(* Logix 5000 project; controller NWGG 1756-L72 rev 35.12; software revision 35.00; part 6 of 19 *)
(* tags used below, declared in another part *)
   _124MB : ALIAS FOR B9[124].2;
   _124STB : ALIAS FOR B9[124].0;
   _124STPB : ALIAS FOR B9[124].1;
   _24_16_0 : ALIAS FOR N250[0];
   _24_16_1 : ALIAS FOR N250[1];
   _24_16_2 : ALIAS FOR N250[2];
   _24_16_3 : ALIAS FOR N250[3];
   _24_16_4 : ALIAS FOR N250[4];
   _24_16_5 : ALIAS FOR N250[5];
   _24_16_6 : ALIAS FOR N250[6];
   _24_16_7 : ALIAS FOR N250[7];
   _24_17_0 : ALIAS FOR N240[0];
   _24_18_0_AN : ALIAS FOR N230[10];
   _24_18_1_AN : ALIAS FOR N230[11];
   _24_18_2_AN : ALIAS FOR N230[12];
   _24_18_3_AN : ALIAS FOR N230[13];
   _24_19_0 : ALIAS FOR N220[10];
   _24_19_1 : ALIAS FOR N220[11];
   _24_19_2 : ALIAS FOR N220[12];
   _24_19_3 : ALIAS FOR N220[13];
   _24_20_0 : ALIAS FOR N210[10];
   _45_AIR_SEQ : ALIAS FOR T4[34];
   _45_SEQ_AIR : ALIAS FOR O12.15;
   _45AUTO : ALIAS FOR B9[45].4;
   _45HAND : ALIAS FOR B9[45].3;
   _45M : ALIAS FOR O25[8].7;
   _45MB : ALIAS FOR B9[45].2;
   _45STB : ALIAS FOR B9[45].0;
   _45STPB : ALIAS FOR B9[45].1;
   _45Y : ALIAS FOR I25[0].7;
   _46AUTO : ALIAS FOR B9[46].4;
   _46HAND : ALIAS FOR B9[46].3;
   _46M : ALIAS FOR O25[8].8;
   _46MB : ALIAS FOR B9[46].2;
   _46STB : ALIAS FOR B9[46].0;
   _46STPB : ALIAS FOR B9[46].1;
   _46Y : ALIAS FOR I25[0].8;
   _47M : ALIAS FOR O25[9].10;
   _47MB : ALIAS FOR B9[47].2;
   _47Y : ALIAS FOR I25[1].10;
   _700_TREAT : ALIAS FOR I7.3;
   _9_TRT_MOV : ALIAS FOR O24[7].4;
   ALARM_FIEL : ALIAS FOR T11[7];
   ALARM_HAND : ALIAS FOR B3[0].10;
   ALARM_HORN : ALIAS FOR O25[11].15;
   ALARM_HORN1 : ALIAS FOR O12.14;
   ALARM_LIGH : ALIAS FOR O13.15;
   ALARM_LT_O : ALIAS FOR T11[3];
   ALARM_SILE : ALIAS FOR I25[4].7;
   ALARM_SILE1 : ALIAS FOR I7.13;
   ALARM_SILE2 : ALIAS FOR B3[0].3;
   ALARM_SILE4 : ALIAS FOR B3[0].9;
   ALRM_LIGHT : ALIAS FOR O25[11].14;
   ALRM_SILEN : ALIAS FOR B3[0].7;
   B3 : DINT[250];
   I24_004_Bit00 : ALIAS FOR I24[4].0;
   I24_004_Bit01 : ALIAS FOR I24[4].1;
   I24_004_Bit02 : ALIAS FOR I24[4].2;
   I24_004_Bit03 : ALIAS FOR I24[4].3;
   I24_004_Bit04 : ALIAS FOR I24[4].4;
   I24_004_Bit05 : ALIAS FOR I24[4].5;
   I24_004_Bit06 : ALIAS FOR I24[4].6;
   I24_004_Bit07 : ALIAS FOR I24[4].7;
   I24_004_Bit08 : ALIAS FOR I24[4].8;
   I24_006_Bit02 : ALIAS FOR I24[6].2;
   I24_021_Bit00 : ALIAS FOR I24[21].0;
   I24_021_Bit01 : ALIAS FOR I24[21].1;
   I24_021_Bit02 : ALIAS FOR I24[21].2;
   I24_021_Bit03 : ALIAS FOR I24[21].3;
   I24_021_Bit04 : ALIAS FOR I24[21].4;
   I24_021_Bit05 : ALIAS FOR I24[21].5;
   I24_021_Bit06 : ALIAS FOR I24[21].6;
   I24_021_Bit07 : ALIAS FOR I24[21].7;
   I24_021_Bit08 : ALIAS FOR I24[21].8;
   IE8_BTR_FL : ALIAS FOR N23[0];
   MAIN_TIMER1 : ALIAS FOR T11[1];
   N23 : DINT[5];
   O24_005_Bit15 : ALIAS FOR O24[5].15;
   O24_007_Bit10 : ALIAS FOR O24[7].10;
   P10_FLOW_A : ALIAS FOR N13[82];
   P10_FLOW_P1 : ALIAS FOR C5[39];
   P10_FLW_OZ : ALIAS FOR N13[80];
   P10_MB : ALIAS FOR B12[10].2;
   P10_OZ : ALIAS FOR N13[81];
   P10_SET : ALIAS FOR B12[10].0;
   P10_SPEED : ALIAS FOR N13[84];
   P10_STOP : ALIAS FOR B12[10].1;
   P1_FLOW_AN : ALIAS FOR N13[2];
   P1_FLOW_PL : ALIAS FOR C5[30];
   P1_FLW_OZ : ALIAS FOR N13[0];
   P1_MB : ALIAS FOR B12[1].2;
   P1_OZ : ALIAS FOR N13[1];
   P1_SET : ALIAS FOR B12[1].0;
   P1_SPEED_O : ALIAS FOR N13[4];
   P1_STOP : ALIAS FOR B12[1].1;
   P2_FLOW_AN : ALIAS FOR N13[12];
   P2_FLOW_PL : ALIAS FOR C5[32];
   P2_FLW_OZ : ALIAS FOR N13[10];
   P2_MB : ALIAS FOR B12[2].2;
   P2_OZ : ALIAS FOR N13[11];
   P2_SET : ALIAS FOR B12[2].0;
   P2_SPEED_O : ALIAS FOR N13[14];
   P2_STOP : ALIAS FOR B12[2].1;
   P3_FLOW_AN : ALIAS FOR N13[22];
   P3_FLOW_PL : ALIAS FOR C5[33];
   P3_FLW_OZ : ALIAS FOR N13[20];
   P3_MB : ALIAS FOR B12[3].2;
   P3_OZ : ALIAS FOR N13[21];
   P3_SET : ALIAS FOR B12[3].0;
   P3_SPEED_O : ALIAS FOR N13[24];
   P3_STOP : ALIAS FOR B12[3].1;
   P4_FLOW_AN : ALIAS FOR N13[32];
   P4_FLOW_PL : ALIAS FOR C5[34];
   P4_FLW_OZ : ALIAS FOR N13[30];
   P4_MB : ALIAS FOR B12[4].2;
   P4_OZ : ALIAS FOR N13[31];
   P4_SET : ALIAS FOR B12[4].0;
   P4_SPEED_O : ALIAS FOR N13[34];
   P4_STOP : ALIAS FOR B12[4].1;
   P5_FLOW_AN : ALIAS FOR N13[42];
   P5_FLOW_PL : ALIAS FOR C5[35];
   P5_FLW_OZ : ALIAS FOR N13[40];
   P5_MB : ALIAS FOR B12[5].2;
   P5_OZ : ALIAS FOR N13[41];
   P5_SET : ALIAS FOR B12[5].0;
   P5_SPEED_O : ALIAS FOR N13[44];
   P5_STOP : ALIAS FOR B12[5].1;
   P6_FLOW_AN : ALIAS FOR N13[52];
   P6_FLOW_PL : ALIAS FOR C5[36];
   P6_FLW_OZ : ALIAS FOR N13[50];
   P6_MB : ALIAS FOR B12[6].2;
   P6_OZ : ALIAS FOR N13[51];
   P6_SET : ALIAS FOR B12[6].0;
   P6_SPEED_O : ALIAS FOR N13[54];
   P6_STOP : ALIAS FOR B12[6].1;
   P7_FLOW_AN : ALIAS FOR N13[62];
   P7_FLOW_PL : ALIAS FOR C5[37];
   P7_FLW_OZ : ALIAS FOR N13[60];
   P7_MB : ALIAS FOR B12[7].2;
   P7_OZ : ALIAS FOR N13[61];
   P7_SET : ALIAS FOR B12[7].0;
   P7_SPEED_O : ALIAS FOR N13[64];
   P7_STOP : ALIAS FOR B12[7].1;
   P8_FLOW_AN : ALIAS FOR N13[72];
   P8_FLOW_PL : ALIAS FOR C5[38];
   P8_FLW_OZ : ALIAS FOR N13[70];
   P8_MB : ALIAS FOR B12[8].2;
   P8_OZ : ALIAS FOR N13[71];
   P8_SET : ALIAS FOR B12[8].0;
   P8_SPEED_O : ALIAS FOR N13[74];
   P8_STOP : ALIAS FOR B12[8].1;
   P_RESET_AU : ALIAS FOR B3[4].0;
   RSVIEW_ALA : ALIAS FOR B3[0].11;
   T11_DLY_TR : ALIAS FOR T4[0].PRE;
   T11_DLY_TR2 : ALIAS FOR T4[1].PRE;
   T11_SET_DE : ALIAS FOR B3[2].0;
   T11_TREAT : ALIAS FOR B3[11].0;
   T11_TRT_MO1 : ALIAS FOR T4[41].PRE;
   T12_DLY_TR1 : ALIAS FOR T4[2].PRE;
   T12_DLY_TR4 : ALIAS FOR T4[3].PRE;
   T12_SET_DE : ALIAS FOR B3[2].1;
   T12_TREAT : ALIAS FOR B3[12].0;
   T12_TRT_MO1 : ALIAS FOR T4[42].PRE;
   T13_DLY_TR1 : ALIAS FOR T4[4].PRE;
   T13_DLY_TR4 : ALIAS FOR T4[5].PRE;
   T13_SET_DE : ALIAS FOR B3[2].2;
   T13_TREAT : ALIAS FOR B3[13].0;
   T13_TRT_MO1 : ALIAS FOR T4[43].PRE;
   T13C_CLOSE1 : ALIAS FOR T22[6].PRE;
   T13C_SET_D : ALIAS FOR B21[70].14;
   T13C_TRT_M1 : ALIAS FOR T22[7].PRE;
   T13C_TRT_O1 : ALIAS FOR T22[5].PRE;
   T14_DLY_TR2 : ALIAS FOR T4[6].ACC;
   T14_DLY_TR4 : ALIAS FOR T4[7].PRE;
   T14_SET_DE : ALIAS FOR B3[2].3;
   T14_TREAT : ALIAS FOR B3[14].0;
   T14_TRT_MO1 : ALIAS FOR T4[44].PRE;
   T15_SET_DE : ALIAS FOR B3[2].4;
   T15_TREAT : ALIAS FOR B3[15].0;
   T15_TRT_MO1 : ALIAS FOR T4[45].PRE;
   T15_TRT_OF1 : ALIAS FOR T4[9].PRE;
   T15_TRT_ON1 : ALIAS FOR T4[8].PRE;
   T16_SET_DE : ALIAS FOR B3[2].5;
   T16_TREAT : ALIAS FOR B3[16].0;
   T16_TRT_MO1 : ALIAS FOR T4[46].PRE;
   T16_TRT_OF1 : ALIAS FOR T4[11].PRE;
   T16_TRT_ON1 : ALIAS FOR T4[10].PRE;
   T17_SET_DE : ALIAS FOR B3[2].6;
   T17_TREAT : ALIAS FOR B3[17].0;
   T17_TRT_MO1 : ALIAS FOR T4[47].PRE;
   T17_TRT_OF1 : ALIAS FOR T4[13].PRE;
   T17_TRT_ON1 : ALIAS FOR T4[12].PRE;
   T19 : TIMER[2];
   T19C_CLOSE2 : ALIAS FOR T22[3].PRE;
   T19C_SET_D : ALIAS FOR B21[71].14;
   T19C_TRT_M1 : ALIAS FOR T22[4].PRE;
   T19C_TRT_O1 : ALIAS FOR T22[0].PRE;
   T21_SET_DE : ALIAS FOR B3[2].7;
   T21_TREAT : ALIAS FOR B3[21].0;
   T21_TRT_MO1 : ALIAS FOR T4[48].PRE;
   T21_TRT_OF1 : ALIAS FOR T4[15].PRE;
   T21_TRT_ON1 : ALIAS FOR T4[14].PRE;
   T22_SET_DE : ALIAS FOR B3[2].8;
   T22_TREAT : ALIAS FOR B3[22].0;
   T22_TRT_MO1 : ALIAS FOR T4[49].PRE;
   T22_TRT_OF1 : ALIAS FOR T4[17].PRE;
   T22_TRT_ON1 : ALIAS FOR T4[16].PRE;
   T23_SET_DE : ALIAS FOR B3[2].9;
   T23_TREAT : ALIAS FOR B3[23].0;
   T23_TRT_MO1 : ALIAS FOR T4[50].PRE;
   T23_TRT_OF1 : ALIAS FOR T4[19].PRE;
   T23_TRT_ON1 : ALIAS FOR T4[18].PRE;
   T24_SET_DE : ALIAS FOR B3[2].10;
   T24_TREAT : ALIAS FOR B3[24].0;
   T24_TRT_MO1 : ALIAS FOR T4[51].PRE;
   T24_TRT_OF1 : ALIAS FOR T4[21].PRE;
   T24_TRT_ON1 : ALIAS FOR T4[20].PRE;
   T25_SET_DE : ALIAS FOR B3[2].11;
   T25_TREAT : ALIAS FOR B3[25].0;
   T25_TRT_MO1 : ALIAS FOR T4[52].PRE;
   T25_TRT_OF1 : ALIAS FOR T4[23].PRE;
   T25_TRT_ON1 : ALIAS FOR T4[22].PRE;
   T26_SET_DE : ALIAS FOR B3[2].12;
   T26_TREAT : ALIAS FOR B3[26].0;
   T26_TRT_MO1 : ALIAS FOR T4[53].PRE;
   T26_TRT_OF1 : ALIAS FOR T4[25].PRE;
   T26_TRT_ON1 : ALIAS FOR T4[24].PRE;
   T27_SET_DE : ALIAS FOR B3[2].13;
   T27_TREAT : ALIAS FOR B3[27].0;
   T27_TRT_MO1 : ALIAS FOR T4[54].PRE;
   T27_TRT_OF1 : ALIAS FOR T4[27].PRE;
   T27_TRT_ON1 : ALIAS FOR T4[26].PRE;
   T28_SET_DE : ALIAS FOR B3[2].14;
   T28_TREAT : ALIAS FOR B3[28].0;
   T28_TRT_MO1 : ALIAS FOR T4[55].PRE;
   T28_TRT_OF1 : ALIAS FOR T4[29].PRE;
   T28_TRT_ON1 : ALIAS FOR T4[28].PRE;
   T29_SET_DE : ALIAS FOR B3[2].15;
   T29_TREAT : ALIAS FOR B3[29].0;
   T29_TRT_MO1 : ALIAS FOR T4[56].PRE;
   T29_TRT_OF1 : ALIAS FOR T4[31].PRE;
   T29_TRT_ON1 : ALIAS FOR T4[30].PRE;
   TRT_PumpRATE : DINT[50];
(* _2_MAIN, continued *)

ROUTINE _10_RAW_MOTORS   (* ladder *)
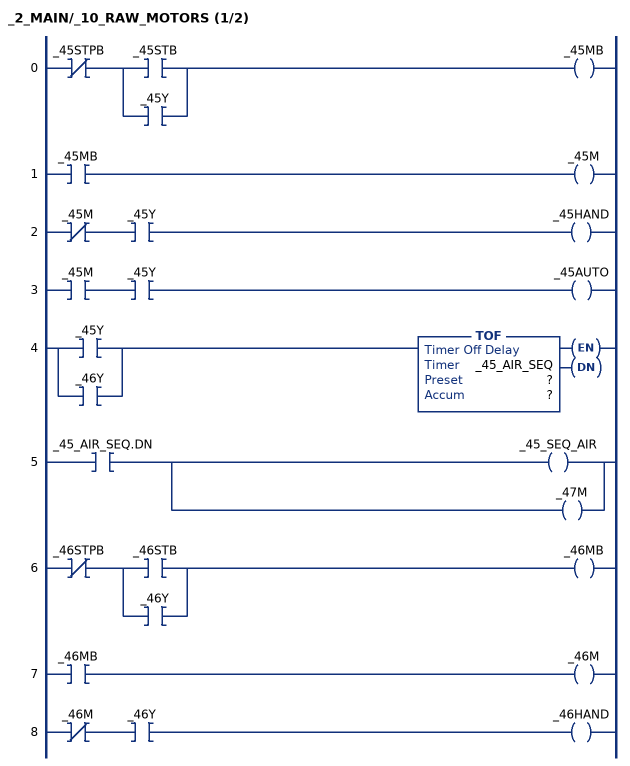
   0: XIO(_45STPB)[XIC(_45STB) ,XIC(_45Y) ]OTE(_45MB);
   1: XIC(_45MB)OTE(_45M);
   2: XIO(_45M)XIC(_45Y)OTE(_45HAND);
   3: XIC(_45M)XIC(_45Y)OTE(_45AUTO);
   4: [XIC(_45Y) ,XIC(_46Y) ]TOF(_45_AIR_SEQ,?,?);
   5: XIC(_45_AIR_SEQ.DN)[OTE(_45_SEQ_AIR) ,OTE(_47M) ];
   6: XIO(_46STPB)[XIC(_46STB) ,XIC(_46Y) ]OTE(_46MB);
   7: XIC(_46MB)OTE(_46M);
   8: XIO(_46M)XIC(_46Y)OTE(_46HAND);
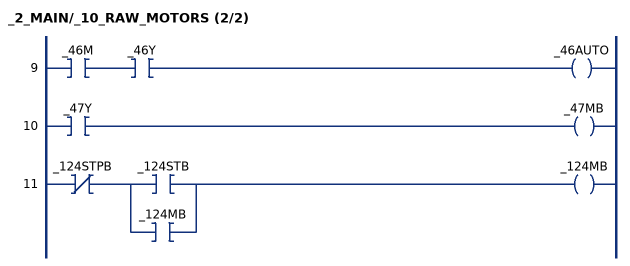
   9: XIC(_46M)XIC(_46Y)OTE(_46AUTO);
   10: XIC(_47Y)OTE(_47MB);
   11: XIO(_124STPB)[XIC(_124STB) ,XIC(_124MB) ]OTE(_124MB);
END_ROUTINE

ROUTINE _34_34_ALARMS   (* ladder *)
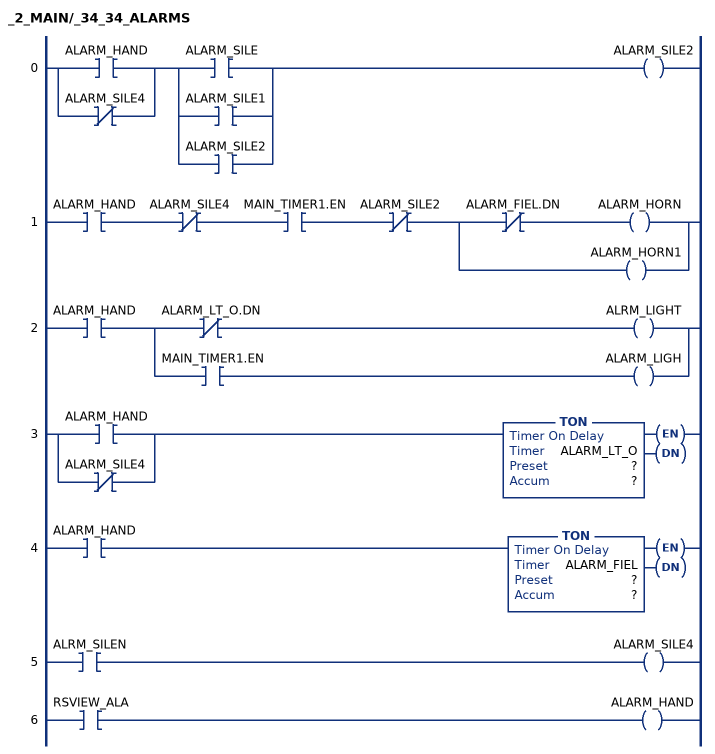
   0: [XIC(ALARM_HAND) ,XIO(ALARM_SILE4) ][XIC(ALARM_SILE) ,XIC(ALARM_SILE1) ,XIC(ALARM_SILE2) ]OTE(ALARM_SILE2);
   1: XIC(ALARM_HAND)XIO(ALARM_SILE4)XIC(MAIN_TIMER1.EN)XIO(ALARM_SILE2)[XIO(ALARM_FIEL.DN) OTE(ALARM_HORN) ,OTE(ALARM_HORN1) ];
   2: XIC(ALARM_HAND)[XIO(ALARM_LT_O.DN) OTE(ALRM_LIGHT) ,XIC(MAIN_TIMER1.EN) OTE(ALARM_LIGH) ];
   3: [XIC(ALARM_HAND) ,XIO(ALARM_SILE4) ]TON(ALARM_LT_O,?,?);
   4: XIC(ALARM_HAND)TON(ALARM_FIEL,?,?);
   5: XIC(ALRM_SILEN)OTE(ALARM_SILE4);
   6: XIC(RSVIEW_ALA)OTE(ALARM_HAND);
END_ROUTINE

ROUTINE _35_35_DEFAULT   (* ladder *)
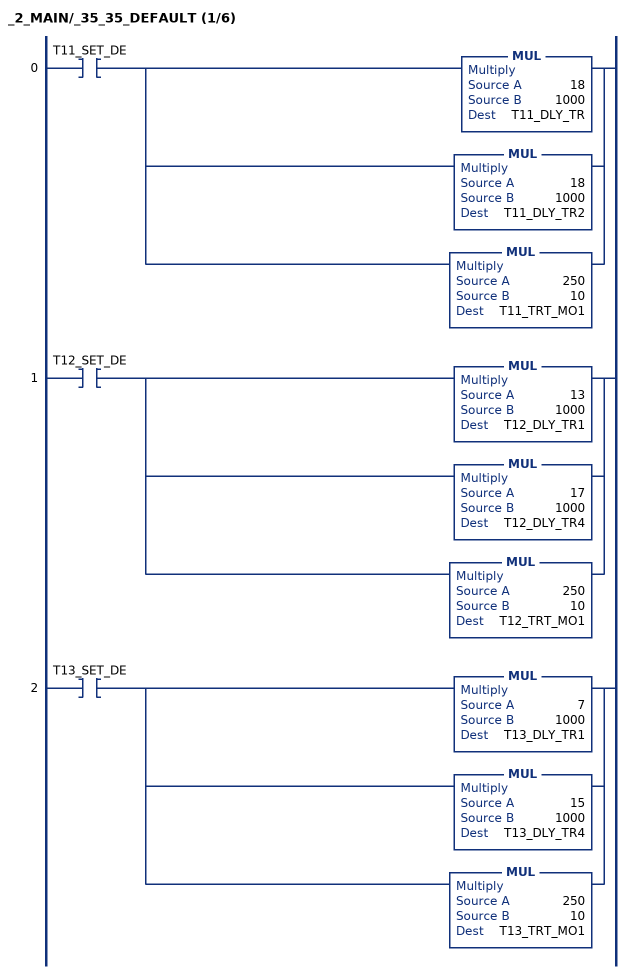
   0: XIC(T11_SET_DE)[MUL(18,1000,T11_DLY_TR) ,MUL(18,1000,T11_DLY_TR2) ,MUL(250,10,T11_TRT_MO1) ];
   1: XIC(T12_SET_DE)[MUL(13,1000,T12_DLY_TR1) ,MUL(17,1000,T12_DLY_TR4) ,MUL(250,10,T12_TRT_MO1) ];
   2: XIC(T13_SET_DE)[MUL(7,1000,T13_DLY_TR1) ,MUL(15,1000,T13_DLY_TR4) ,MUL(250,10,T13_TRT_MO1) ];
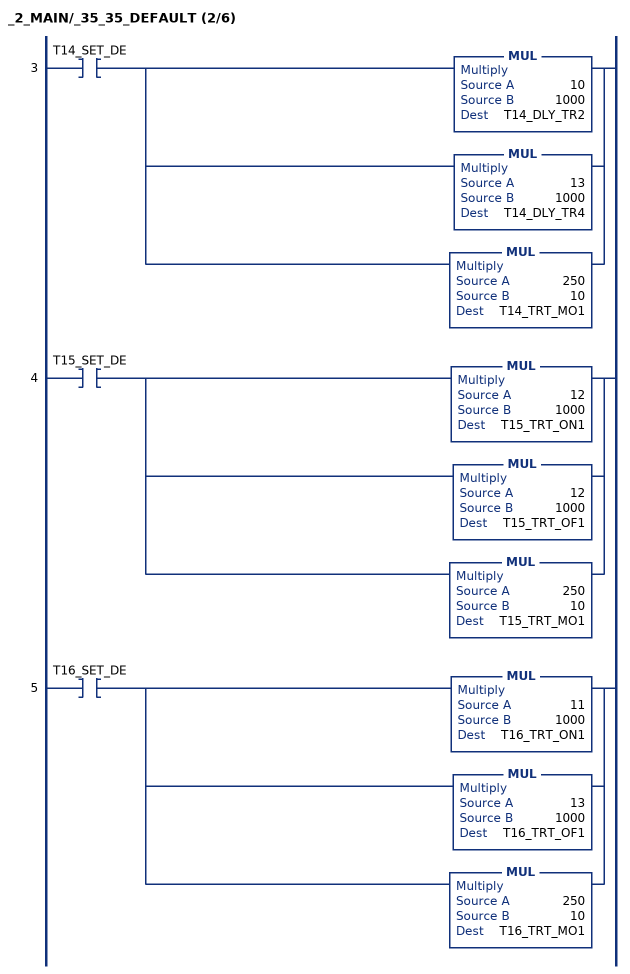
   3: XIC(T14_SET_DE)[MUL(10,1000,T14_DLY_TR2) ,MUL(13,1000,T14_DLY_TR4) ,MUL(250,10,T14_TRT_MO1) ];
   4: XIC(T15_SET_DE)[MUL(12,1000,T15_TRT_ON1) ,MUL(12,1000,T15_TRT_OF1) ,MUL(250,10,T15_TRT_MO1) ];
   5: XIC(T16_SET_DE)[MUL(11,1000,T16_TRT_ON1) ,MUL(13,1000,T16_TRT_OF1) ,MUL(250,10,T16_TRT_MO1) ];
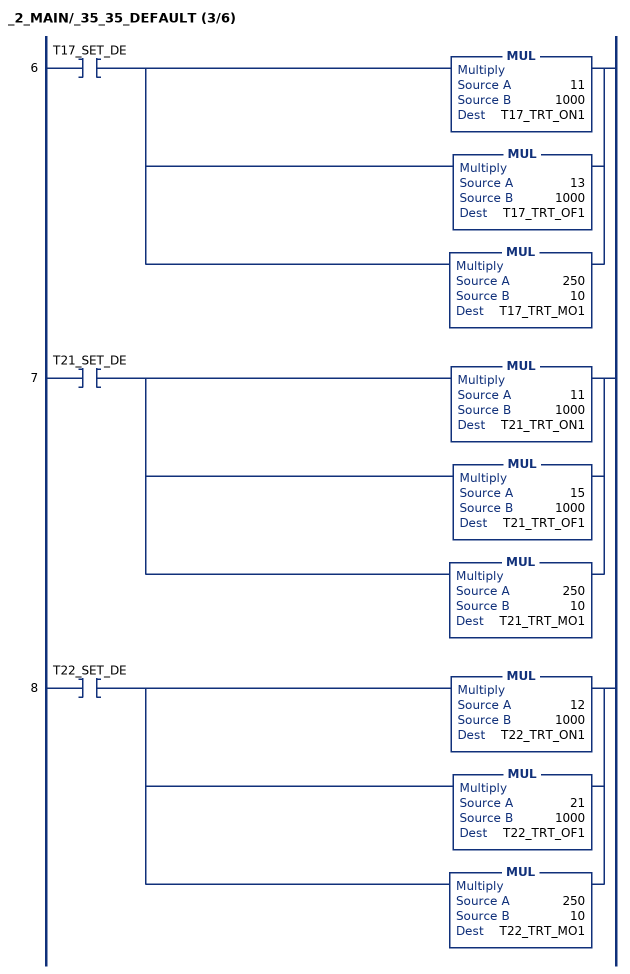
   6: XIC(T17_SET_DE)[MUL(11,1000,T17_TRT_ON1) ,MUL(13,1000,T17_TRT_OF1) ,MUL(250,10,T17_TRT_MO1) ];
   7: XIC(T21_SET_DE)[MUL(11,1000,T21_TRT_ON1) ,MUL(15,1000,T21_TRT_OF1) ,MUL(250,10,T21_TRT_MO1) ];
   8: XIC(T22_SET_DE)[MUL(12,1000,T22_TRT_ON1) ,MUL(21,1000,T22_TRT_OF1) ,MUL(250,10,T22_TRT_MO1) ];
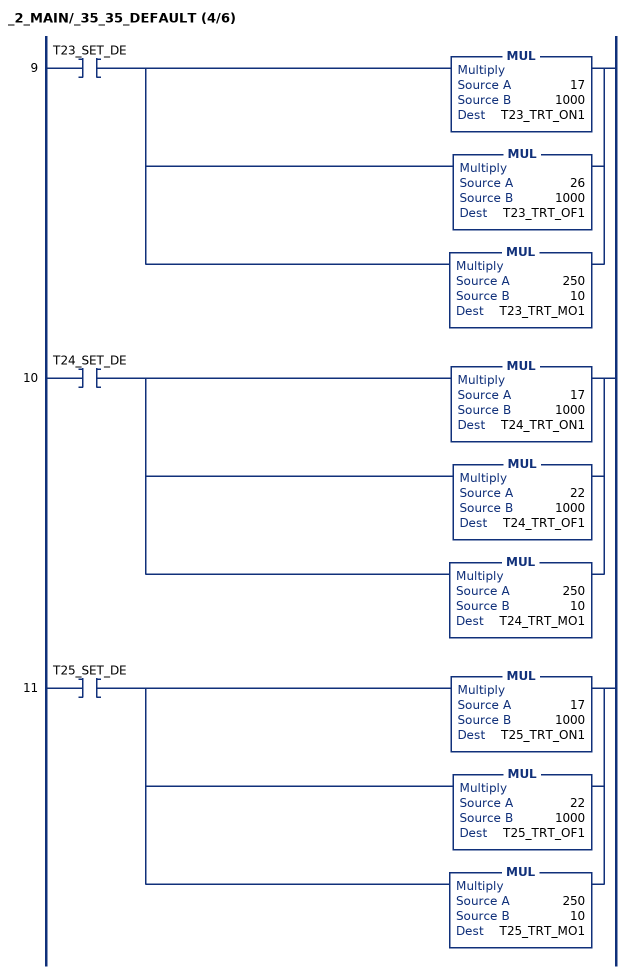
   9: XIC(T23_SET_DE)[MUL(17,1000,T23_TRT_ON1) ,MUL(26,1000,T23_TRT_OF1) ,MUL(250,10,T23_TRT_MO1) ];
   10: XIC(T24_SET_DE)[MUL(17,1000,T24_TRT_ON1) ,MUL(22,1000,T24_TRT_OF1) ,MUL(250,10,T24_TRT_MO1) ];
   11: XIC(T25_SET_DE)[MUL(17,1000,T25_TRT_ON1) ,MUL(22,1000,T25_TRT_OF1) ,MUL(250,10,T25_TRT_MO1) ];
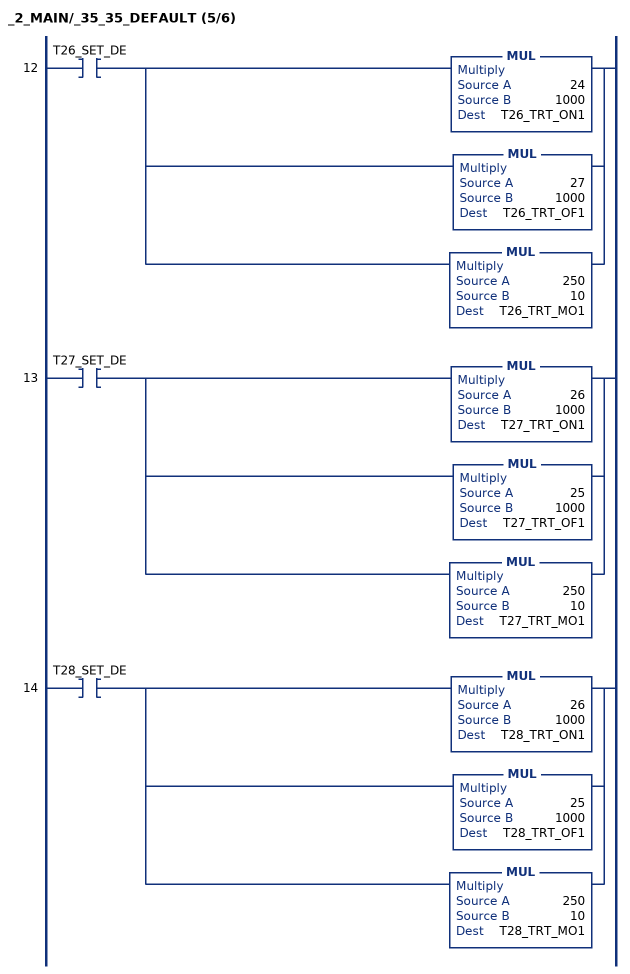
   12: XIC(T26_SET_DE)[MUL(24,1000,T26_TRT_ON1) ,MUL(27,1000,T26_TRT_OF1) ,MUL(250,10,T26_TRT_MO1) ];
   13: XIC(T27_SET_DE)[MUL(26,1000,T27_TRT_ON1) ,MUL(25,1000,T27_TRT_OF1) ,MUL(250,10,T27_TRT_MO1) ];
   14: XIC(T28_SET_DE)[MUL(26,1000,T28_TRT_ON1) ,MUL(25,1000,T28_TRT_OF1) ,MUL(250,10,T28_TRT_MO1) ];
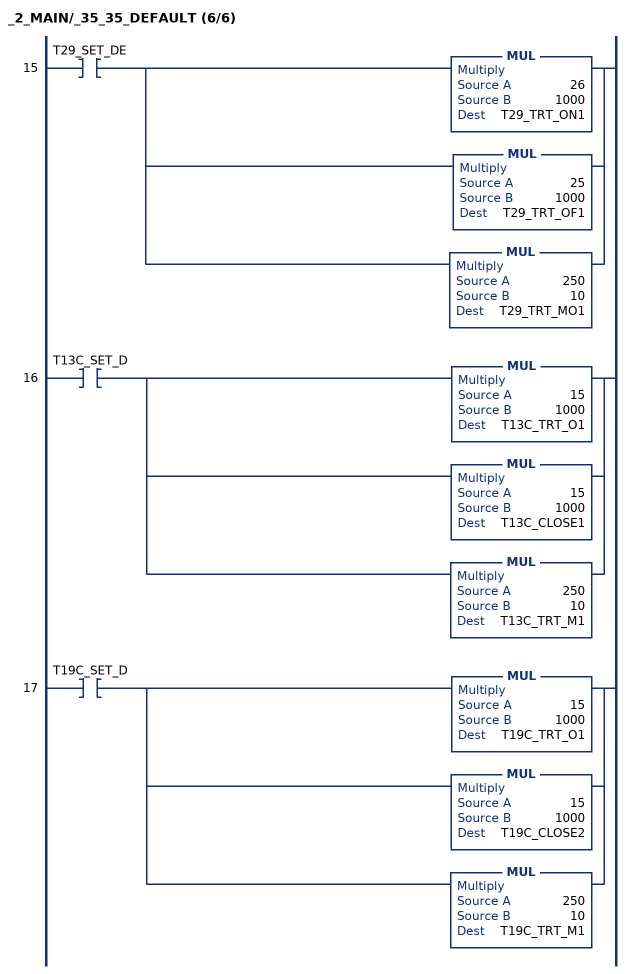
   15: XIC(T29_SET_DE)[MUL(26,1000,T29_TRT_ON1) ,MUL(25,1000,T29_TRT_OF1) ,MUL(250,10,T29_TRT_MO1) ];
   16: XIC(T13C_SET_D)[MUL(15,1000,T13C_TRT_O1) ,MUL(15,1000,T13C_CLOSE1) ,MUL(250,10,T13C_TRT_M1) ];
   17: XIC(T19C_SET_D)[MUL(15,1000,T19C_TRT_O1) ,MUL(15,1000,T19C_CLOSE2) ,MUL(250,10,T19C_TRT_M1) ];
END_ROUTINE

ROUTINE _36_36_TREATER_FLOW_PUMPS   (* ladder *)
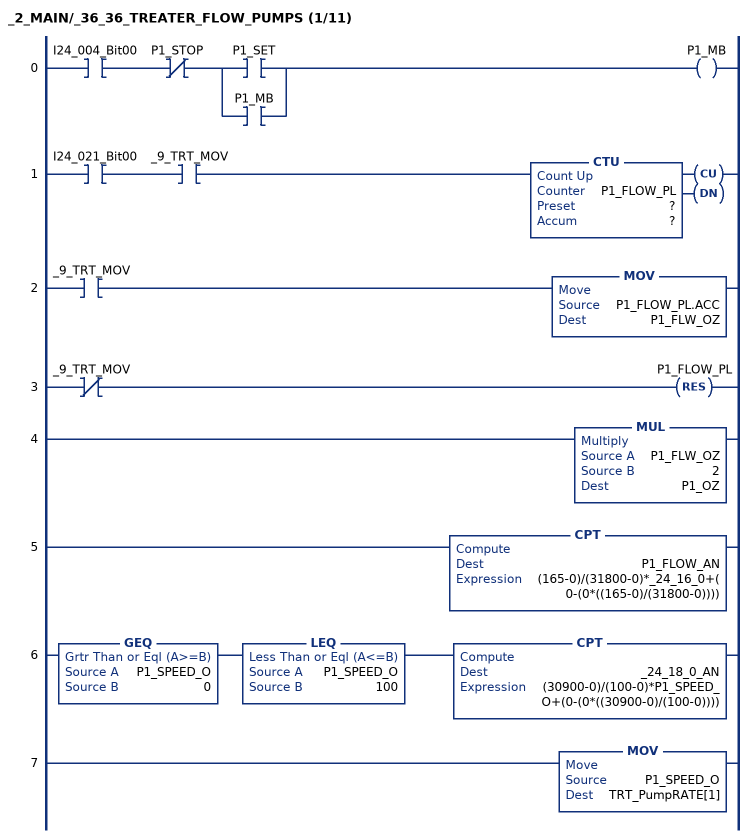
   0: XIC(I24_004_Bit00)XIO(P1_STOP)[XIC(P1_SET) ,XIC(P1_MB) ]OTE(P1_MB);
   1: XIC(I24_021_Bit00)XIC(_9_TRT_MOV)CTU(P1_FLOW_PL,?,?);
   2: XIC(_9_TRT_MOV)MOV(P1_FLOW_PL.ACC,P1_FLW_OZ);
   3: XIO(_9_TRT_MOV)RES(P1_FLOW_PL);
   4: MUL(P1_FLW_OZ,2,P1_OZ);
   5: CPT(P1_FLOW_AN,(165-0)/(31800-0)*_24_16_0+(0-(0*((165-0)/(31800-0)))));
   6: GEQ(P1_SPEED_O,0)LEQ(P1_SPEED_O,100)CPT(_24_18_0_AN,(30900-0)/(100-0)*P1_SPEED_O+(0-(0*((30900-0)/(100-0)))));
   7: MOV(P1_SPEED_O,TRT_PumpRATE[1]);
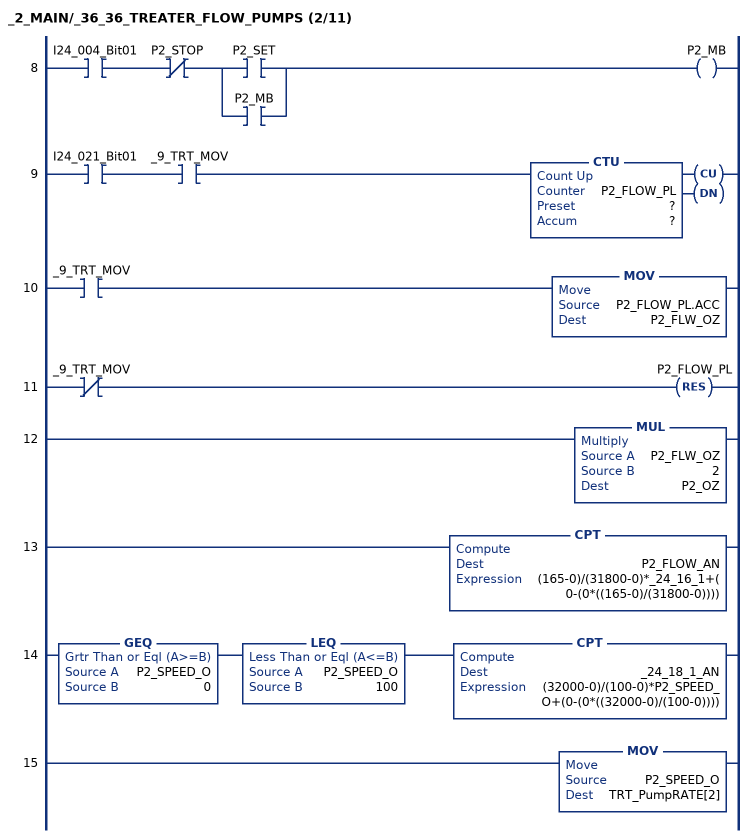
   8: XIC(I24_004_Bit01)XIO(P2_STOP)[XIC(P2_SET) ,XIC(P2_MB) ]OTE(P2_MB);
   9: XIC(I24_021_Bit01)XIC(_9_TRT_MOV)CTU(P2_FLOW_PL,?,?);
   10: XIC(_9_TRT_MOV)MOV(P2_FLOW_PL.ACC,P2_FLW_OZ);
   11: XIO(_9_TRT_MOV)RES(P2_FLOW_PL);
   12: MUL(P2_FLW_OZ,2,P2_OZ);
   13: CPT(P2_FLOW_AN,(165-0)/(31800-0)*_24_16_1+(0-(0*((165-0)/(31800-0)))));
   14: GEQ(P2_SPEED_O,0)LEQ(P2_SPEED_O,100)CPT(_24_18_1_AN,(32000-0)/(100-0)*P2_SPEED_O+(0-(0*((32000-0)/(100-0)))));
   15: MOV(P2_SPEED_O,TRT_PumpRATE[2]);
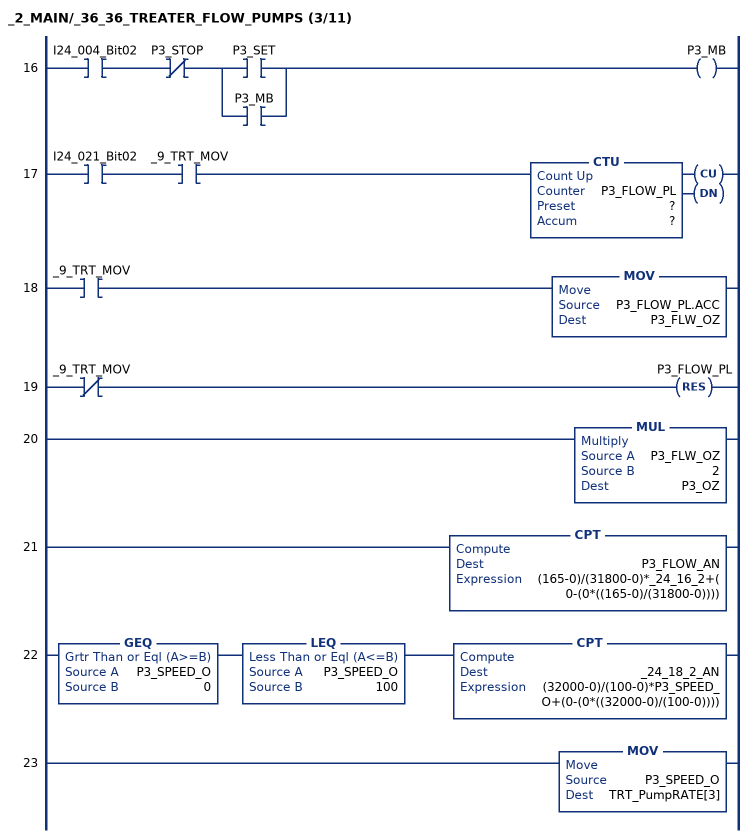
   16: XIC(I24_004_Bit02)XIO(P3_STOP)[XIC(P3_SET) ,XIC(P3_MB) ]OTE(P3_MB);
   17: XIC(I24_021_Bit02)XIC(_9_TRT_MOV)CTU(P3_FLOW_PL,?,?);
   18: XIC(_9_TRT_MOV)MOV(P3_FLOW_PL.ACC,P3_FLW_OZ);
   19: XIO(_9_TRT_MOV)RES(P3_FLOW_PL);
   20: MUL(P3_FLW_OZ,2,P3_OZ);
   21: CPT(P3_FLOW_AN,(165-0)/(31800-0)*_24_16_2+(0-(0*((165-0)/(31800-0)))));
   22: GEQ(P3_SPEED_O,0)LEQ(P3_SPEED_O,100)CPT(_24_18_2_AN,(32000-0)/(100-0)*P3_SPEED_O+(0-(0*((32000-0)/(100-0)))));
   23: MOV(P3_SPEED_O,TRT_PumpRATE[3]);
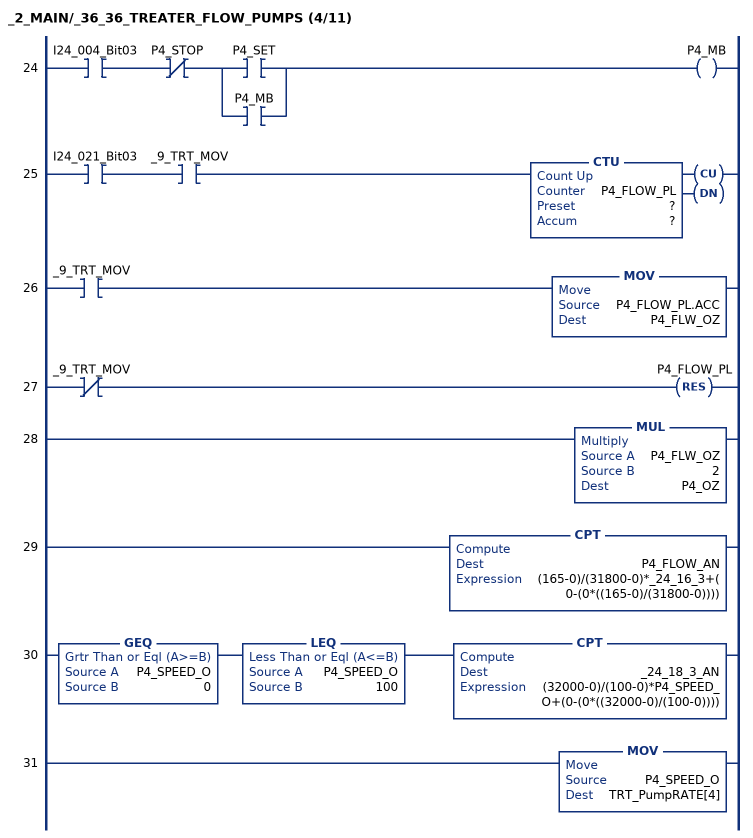
   24: XIC(I24_004_Bit03)XIO(P4_STOP)[XIC(P4_SET) ,XIC(P4_MB) ]OTE(P4_MB);
   25: XIC(I24_021_Bit03)XIC(_9_TRT_MOV)CTU(P4_FLOW_PL,?,?);
   26: XIC(_9_TRT_MOV)MOV(P4_FLOW_PL.ACC,P4_FLW_OZ);
   27: XIO(_9_TRT_MOV)RES(P4_FLOW_PL);
   28: MUL(P4_FLW_OZ,2,P4_OZ);
   29: CPT(P4_FLOW_AN,(165-0)/(31800-0)*_24_16_3+(0-(0*((165-0)/(31800-0)))));
   30: GEQ(P4_SPEED_O,0)LEQ(P4_SPEED_O,100)CPT(_24_18_3_AN,(32000-0)/(100-0)*P4_SPEED_O+(0-(0*((32000-0)/(100-0)))));
   31: MOV(P4_SPEED_O,TRT_PumpRATE[4]);
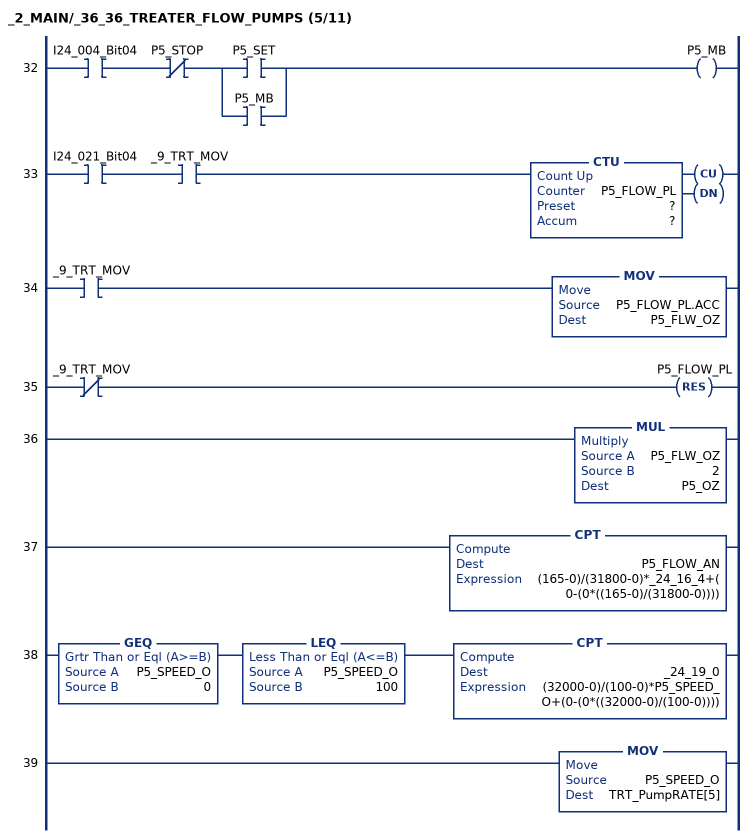
   32: XIC(I24_004_Bit04)XIO(P5_STOP)[XIC(P5_SET) ,XIC(P5_MB) ]OTE(P5_MB);
   33: XIC(I24_021_Bit04)XIC(_9_TRT_MOV)CTU(P5_FLOW_PL,?,?);
   34: XIC(_9_TRT_MOV)MOV(P5_FLOW_PL.ACC,P5_FLW_OZ);
   35: XIO(_9_TRT_MOV)RES(P5_FLOW_PL);
   36: MUL(P5_FLW_OZ,2,P5_OZ);
   37: CPT(P5_FLOW_AN,(165-0)/(31800-0)*_24_16_4+(0-(0*((165-0)/(31800-0)))));
   38: GEQ(P5_SPEED_O,0)LEQ(P5_SPEED_O,100)CPT(_24_19_0,(32000-0)/(100-0)*P5_SPEED_O+(0-(0*((32000-0)/(100-0)))));
   39: MOV(P5_SPEED_O,TRT_PumpRATE[5]);
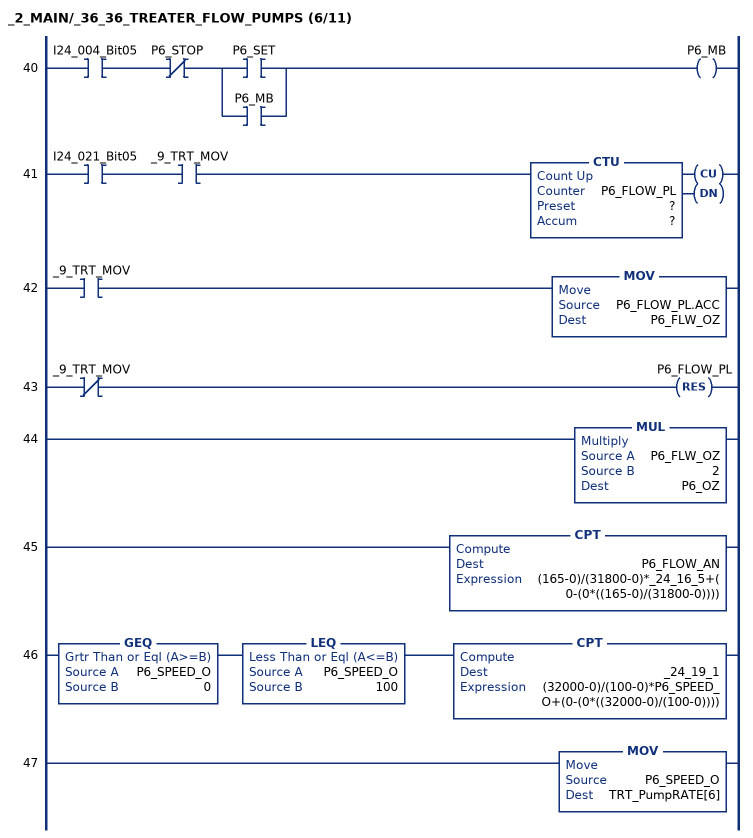
   40: XIC(I24_004_Bit05)XIO(P6_STOP)[XIC(P6_SET) ,XIC(P6_MB) ]OTE(P6_MB);
   41: XIC(I24_021_Bit05)XIC(_9_TRT_MOV)CTU(P6_FLOW_PL,?,?);
   42: XIC(_9_TRT_MOV)MOV(P6_FLOW_PL.ACC,P6_FLW_OZ);
   43: XIO(_9_TRT_MOV)RES(P6_FLOW_PL);
   44: MUL(P6_FLW_OZ,2,P6_OZ);
   45: CPT(P6_FLOW_AN,(165-0)/(31800-0)*_24_16_5+(0-(0*((165-0)/(31800-0)))));
   46: GEQ(P6_SPEED_O,0)LEQ(P6_SPEED_O,100)CPT(_24_19_1,(32000-0)/(100-0)*P6_SPEED_O+(0-(0*((32000-0)/(100-0)))));
   47: MOV(P6_SPEED_O,TRT_PumpRATE[6]);
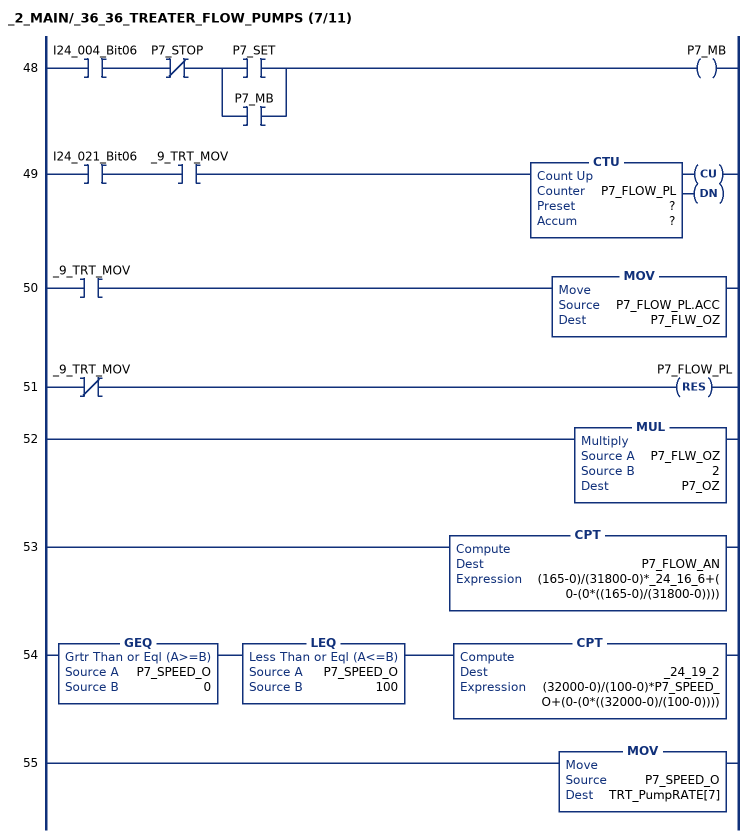
   48: XIC(I24_004_Bit06)XIO(P7_STOP)[XIC(P7_SET) ,XIC(P7_MB) ]OTE(P7_MB);
   49: XIC(I24_021_Bit06)XIC(_9_TRT_MOV)CTU(P7_FLOW_PL,?,?);
   50: XIC(_9_TRT_MOV)MOV(P7_FLOW_PL.ACC,P7_FLW_OZ);
   51: XIO(_9_TRT_MOV)RES(P7_FLOW_PL);
   52: MUL(P7_FLW_OZ,2,P7_OZ);
   53: CPT(P7_FLOW_AN,(165-0)/(31800-0)*_24_16_6+(0-(0*((165-0)/(31800-0)))));
   54: GEQ(P7_SPEED_O,0)LEQ(P7_SPEED_O,100)CPT(_24_19_2,(32000-0)/(100-0)*P7_SPEED_O+(0-(0*((32000-0)/(100-0)))));
   55: MOV(P7_SPEED_O,TRT_PumpRATE[7]);
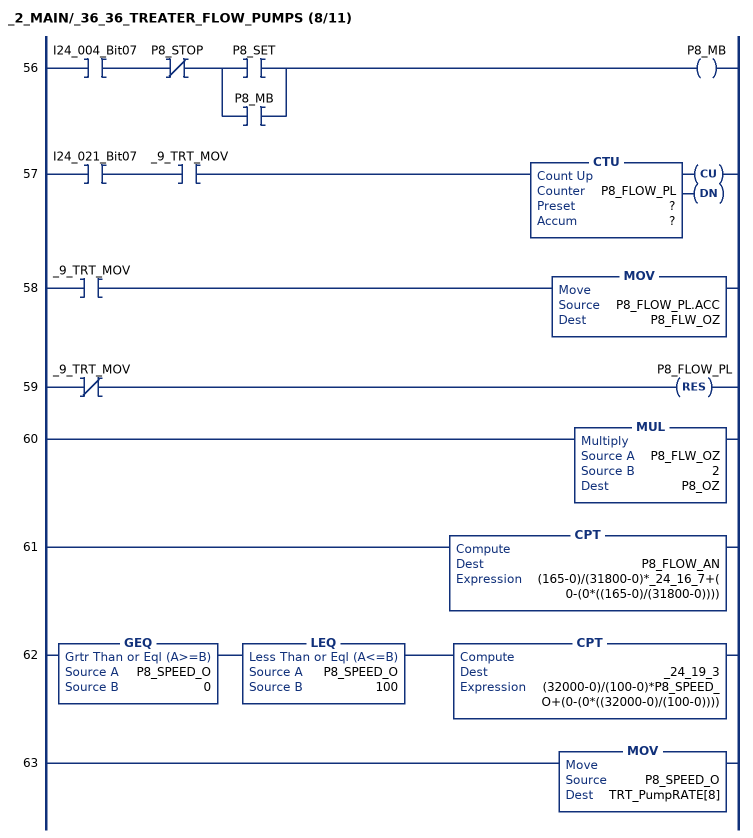
   56: XIC(I24_004_Bit07)XIO(P8_STOP)[XIC(P8_SET) ,XIC(P8_MB) ]OTE(P8_MB);
   57: XIC(I24_021_Bit07)XIC(_9_TRT_MOV)CTU(P8_FLOW_PL,?,?);
   58: XIC(_9_TRT_MOV)MOV(P8_FLOW_PL.ACC,P8_FLW_OZ);
   59: XIO(_9_TRT_MOV)RES(P8_FLOW_PL);
   60: MUL(P8_FLW_OZ,2,P8_OZ);
   61: CPT(P8_FLOW_AN,(165-0)/(31800-0)*_24_16_7+(0-(0*((165-0)/(31800-0)))));
   62: GEQ(P8_SPEED_O,0)LEQ(P8_SPEED_O,100)CPT(_24_19_3,(32000-0)/(100-0)*P8_SPEED_O+(0-(0*((32000-0)/(100-0)))));
   63: MOV(P8_SPEED_O,TRT_PumpRATE[8]);
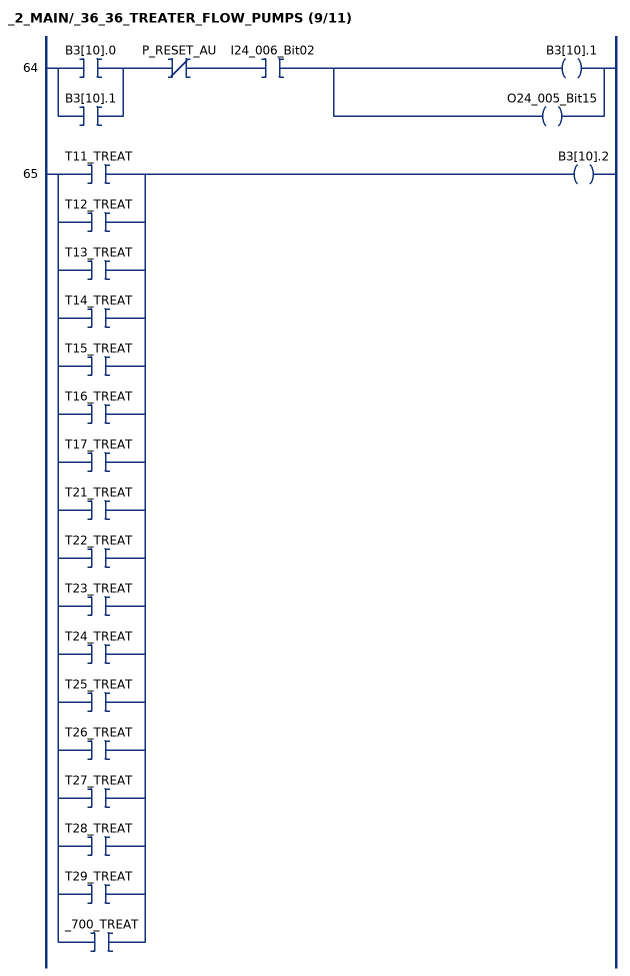
   64: [XIC(B3[10].0) ,XIC(B3[10].1) ]XIO(P_RESET_AU)XIC(I24_006_Bit02)[OTE(B3[10].1) ,OTE(O24_005_Bit15) ];
   65: [XIC(T11_TREAT) ,XIC(T12_TREAT) ,XIC(T13_TREAT) ,XIC(T14_TREAT) ,XIC(T15_TREAT) ,XIC(T16_TREAT) ,XIC(T17_TREAT) ,XIC(T21_TREAT) ,XIC(T22_TREAT) ,XIC(T23_TREAT) ,XIC(T24_TREAT) ,XIC(T25_TREAT) ,XIC(T26_TREAT) ,XIC(T27_TREAT) ,XIC(T28_TREAT) ,XIC(T29_TREAT) ,XIC(_700_TREAT) ]OTE(B3[10].2);
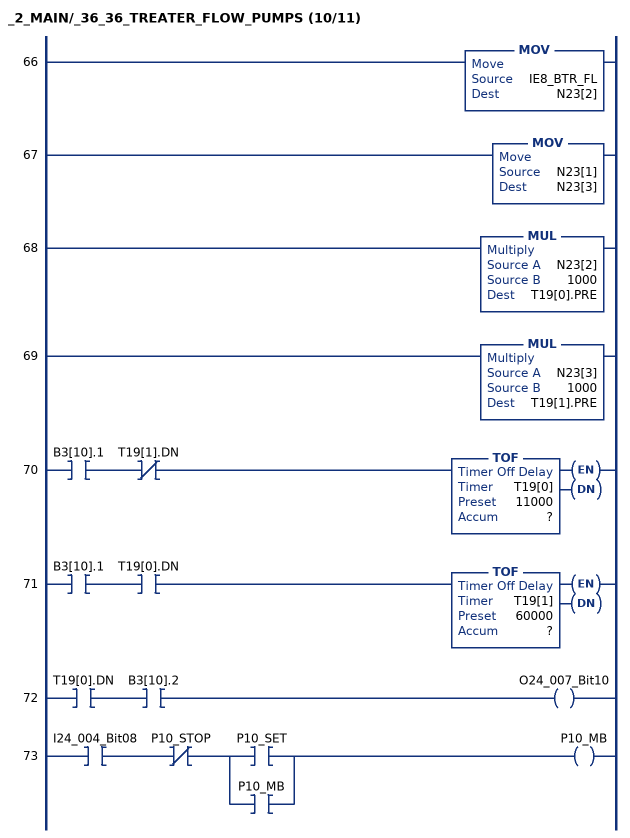
   66: MOV(IE8_BTR_FL,N23[2]);
   67: MOV(N23[1],N23[3]);
   68: MUL(N23[2],1000,T19[0].PRE);
   69: MUL(N23[3],1000,T19[1].PRE);
   70: XIC(B3[10].1)XIO(T19[1].DN)TOF(T19[0],?,?);
   71: XIC(B3[10].1)XIC(T19[0].DN)TOF(T19[1],?,?);
   72: XIC(T19[0].DN)XIC(B3[10].2)OTE(O24_007_Bit10);
   73: XIC(I24_004_Bit08)XIO(P10_STOP)[XIC(P10_SET) ,XIC(P10_MB) ]OTE(P10_MB);
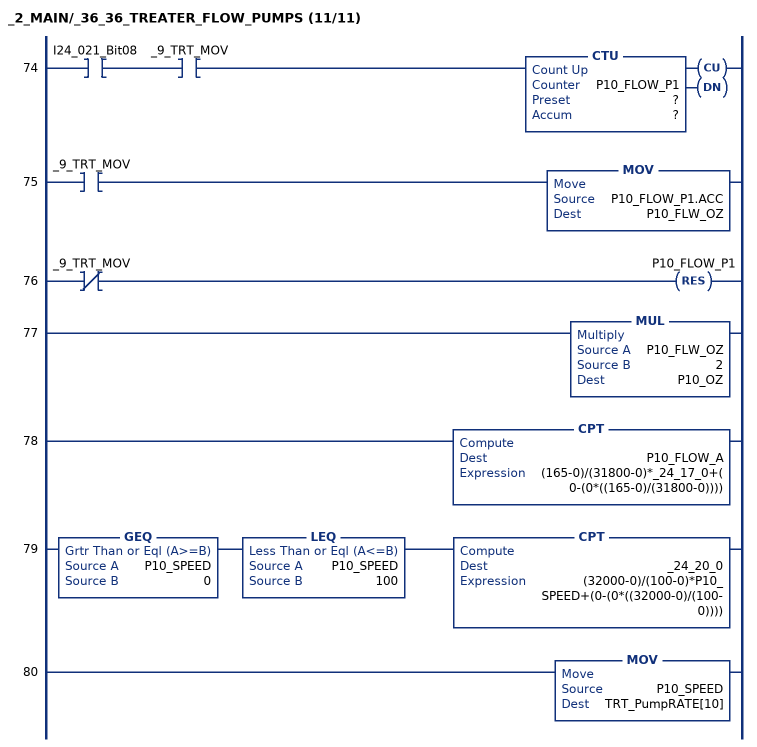
   74: XIC(I24_021_Bit08)XIC(_9_TRT_MOV)CTU(P10_FLOW_P1,?,?);
   75: XIC(_9_TRT_MOV)MOV(P10_FLOW_P1.ACC,P10_FLW_OZ);
   76: XIO(_9_TRT_MOV)RES(P10_FLOW_P1);
   77: MUL(P10_FLW_OZ,2,P10_OZ);
   78: CPT(P10_FLOW_A,(165-0)/(31800-0)*_24_17_0+(0-(0*((165-0)/(31800-0)))));
   79: GEQ(P10_SPEED,0)LEQ(P10_SPEED,100)CPT(_24_20_0,(32000-0)/(100-0)*P10_SPEED+(0-(0*((32000-0)/(100-0)))));
   80: MOV(P10_SPEED,TRT_PumpRATE[10]);
END_ROUTINE
